// TIA Portal project "Est_clasificacion" (V17)

(* hardware
DEVICE "Estación S7-1500/ET200MP_1"  S7-1500 station
   slot 0: "Perfil soporte_0"  Rack  6ES7 590-1***0-0AA0
   slot 1: "PLC_1"  CPU 1516-3 PN/DP  6ES7 516-3AN02-0AB0  V2.9
      slot 3: "Display de la CPU_1"  6ES7591-1BA00-0AA0
      slot 32768: "Interfaz PROFINET_1"  X1
         slot 32769: "Puerto_1"  X1 P1
         slot 32770: "Puerto_2"  X1 P2
      slot 33024: "Interfaz PROFINET_2"  X2
         slot 33025: "Puerto_1"  X2 P1
      slot 33280: "Interfaz DP_1"  X3
      slot 34817: "Virtual CP interface port_1"  Virtual CP interface port  Virtual CP interface port
   slot 2: "DI 32x24VDC HF_1"  DI 32x24VDC HF  6ES7 521-1BL00-0AB0  V2.2
   slot 3: "DQ 32x24VDC/0.5A HF_1"  DQ 32x24VDC/0.5A HF  6ES7 522-1BL01-0AB0  V1.1
   slot 4: "AI 8xU/I/RTD/TC ST_1"  AI 8xU/I/RTD/TC ST  6ES7 531-7KF00-0AB0  V2.2
   slot 5: "AQ 4xU/I ST_1"  AQ 4xU/I ST  6ES7 532-5HD00-0AB0  V2.2
DEVICE "HMI_1"  KTP600 Basic color PN
   slot 0: "HMI_1"  KTP600 Basic color PN  6AV6 647-0AD11-3AX0  12.0.0.0
   slot 1: "HMI_RT_1"  KTP600 Basic color PN  6AV6 647-0AD11-3AX0  12.0.0.0
   slot 5: "HMI_1.IE_CP_1"  PROFINET Interface  12.0.0.0
      slot 1: "Interfaz PROFINET_1"  PROFINET Interface
         slot 1: "Port_1"  Port
*)

// ===== PLC "PLC_1"  CPU 1516-3 PN/DP =====

VAR_GLOBAL   // PLC tag table "Tabla de variables estándar"
   "Detector pieza inicio" AT %I0.0 : Bool;
   "Deflector 1" AT %I0.1 : Bool;
   "Detector de pieza" AT %I0.2 : Bool;
   "Deflector 2" AT %I0.3 : Bool;
   "Detector pieza color" AT %I0.4 : Bool;
   "Detector pieza negra" AT %I0.5 : Bool;
   "Detector pieza metalica" AT %I0.6 : Bool;
   "Start" AT %I1.0 : Bool;
   "Reset" AT %I1.3 : Bool;
   "Avanzar cinta" AT %Q0.0 : Bool;
   "Avanzar deflector 1" AT %Q0.1 : Bool;
   "Avanzar deflector 2" AT %Q0.2 : Bool;
   "Retraer tope" AT %Q0.3 : Bool;
   "Luz ON" AT %Q1.0 : Bool;
   "Luz RESET" AT %Q1.1 : Bool;
   "M0.0" AT %M0.0 : Bool;
   "M0.1" AT %M0.1 : Bool;
   "M0.2" AT %M0.2 : Bool;
   "C0.0" AT %M0.3 : Bool;
   "C0.1" AT %M0.4 : Bool;
   "C0.2" AT %M0.5 : Bool;
   "M1.0" AT %M1.0 : Bool;
   "M1.1" AT %M1.1 : Bool;
   "M1.2" AT %M1.2 : Bool;
   "M1.3" AT %M1.3 : Bool;
   "M1.4" AT %M1.4 : Bool;
   "M1.5" AT %M1.5 : Bool;
   "System_Byte" AT %MB7789 : Byte;
   "FirstScan" AT %M7789.0 : Bool;
   "DiagStatusUpdate" AT %M7789.1 : Bool;
   "AlwaysTRUE" AT %M7789.2 : Bool;
   "AlwaysFALSE" AT %M7789.3 : Bool;
END_VAR

// folder: System blocks/Program resources

DATA_BLOCK "IEC_Timer_0_DB"   // DB1
{ S7_Optimized_Access := 'TRUE' }
AUTHOR : Simatic
FAMILY : IEC
NAME : IEC_TMR
VERSION : 1.0
// stored: InstanceOfName IEC_TIMER
"IEC_TIMER"
BEGIN
END_DATA_BLOCK

DATA_BLOCK "IEC_Counter_0_DB"   // DB4
{ S7_Optimized_Access := 'TRUE' }
AUTHOR : Simatic
FAMILY : IEC
NAME : CNTR
VERSION : 1.0
// stored: InstanceOfName IEC_COUNTER
"IEC_COUNTER"
BEGIN
END_DATA_BLOCK

DATA_BLOCK "IEC_Counter_0_DB_1"   // DB5
{ S7_Optimized_Access := 'TRUE' }
AUTHOR : Simatic
FAMILY : IEC
NAME : CNTR
VERSION : 1.0
// stored: InstanceOfName IEC_COUNTER
"IEC_COUNTER"
BEGIN
END_DATA_BLOCK

DATA_BLOCK "IEC_Counter_0_DB_2"   // DB6
{ S7_Optimized_Access := 'TRUE' }
AUTHOR : Simatic
FAMILY : IEC
NAME : CNTR
VERSION : 1.0
// stored: InstanceOfName IEC_COUNTER
"IEC_COUNTER"
BEGIN
END_DATA_BLOCK

// folder: (top level)

ORGANIZATION_BLOCK "Main"   // OB1, LAD, ProgramCycle
TITLE = "Main Program Sweep (Cycle)"
{ S7_Optimized_Access := 'TRUE' }
VERSION : 0.1
   VAR_INPUT
      Initial_Call : Bool;   // Initial call of this OB
      Remanence : Bool;   // =True, if remanent data are available
   END_VAR
   VAR_TEMP   // added for the SCL form of the ladder/FBD networks
      _w1 : Bool;
      _w2 : Bool;
   END_VAR
BEGIN

REGION Network 1: Estados panel
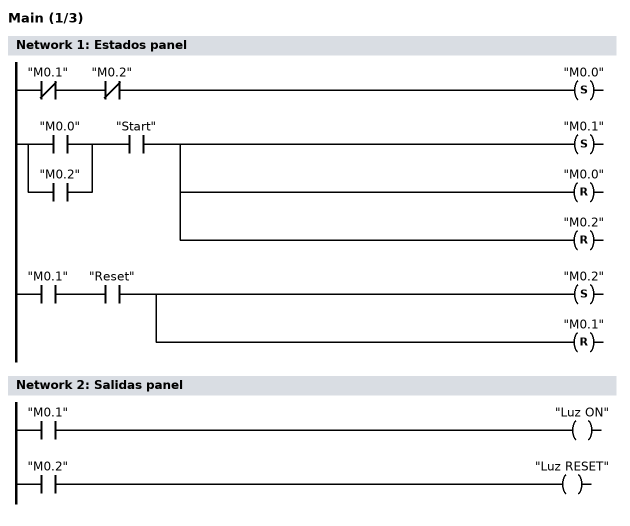
   RUNG wire#powerrail
      I_Contact( "M0.1" )
      I_Contact( "M0.2" )
      S_Coil( "M0.0" )
   END_RUNG
   RUNG wire#powerrail
      Contact( "M0.0" )
      wire#w1
      Contact( "Start" )
      wire#w2
      S_Coil( "M0.1" )
   END_RUNG
   RUNG wire#powerrail
      Contact( "M0.2" )
   END_RUNG wire#w1
   RUNG wire#w2
      R_Coil( "M0.0" )
   END_RUNG
   RUNG wire#w2
      R_Coil( "M0.2" )
   END_RUNG
   RUNG wire#powerrail
      Contact( "M0.1" )
      Contact( "Reset" )
      wire#w3
      S_Coil( "M0.2" )
   END_RUNG
   RUNG wire#w3
      R_Coil( "M0.1" )
   END_RUNG
   // the same network as SCL:
   IF NOT "M0.1" AND NOT "M0.2" THEN "M0.0" := TRUE; END_IF;
   IF ("M0.0" OR "M0.2") AND "Start" THEN "M0.1" := TRUE; END_IF;
   #_w1 := ("M0.0" OR "M0.2") AND "Start";
   IF #_w1 THEN
       "M0.0" := FALSE;
       "M0.2" := FALSE;
   END_IF;
   IF "M0.1" AND "Reset" THEN
       "M0.2" := TRUE;
       "M0.1" := FALSE;
   END_IF;
END_REGION

REGION Network 2: Salidas panel
   RUNG wire#powerrail
      Contact( "M0.1" )
      Coil( "Luz ON" )
   END_RUNG
   RUNG wire#powerrail
      Contact( "M0.2" )
      Coil( "Luz RESET" )
   END_RUNG
   // the same network as SCL:
   "Luz ON" := "M0.1";
   "Luz RESET" := "M0.2";
END_REGION

REGION Network 3: Estados principal
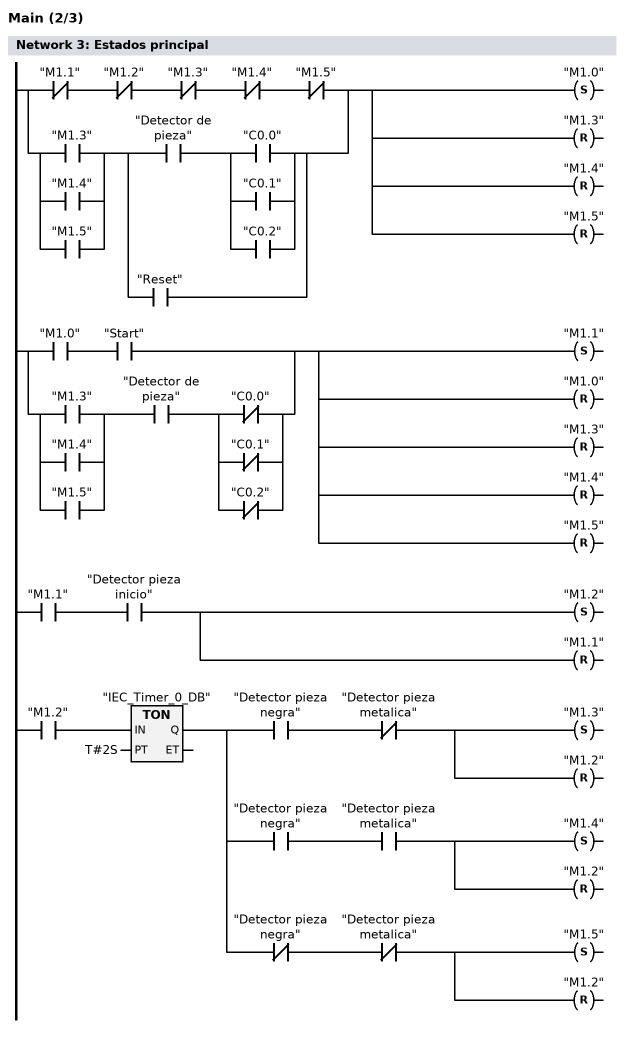
   IF (NOT "M1.1" AND NOT "M1.2" AND NOT "M1.3" AND NOT "M1.4" AND NOT "M1.5") OR (("M1.3" OR "M1.4" OR "M1.5") AND (("Detector de pieza" AND ("C0.0" OR "C0.1" OR "C0.2")) OR "Reset")) THEN
       "M1.0" := TRUE;
   END_IF;
   #_w1 := (NOT "M1.1" AND NOT "M1.2" AND NOT "M1.3" AND NOT "M1.4" AND NOT "M1.5") OR (("M1.3" OR "M1.4" OR "M1.5") AND (("Detector de pieza" AND ("C0.0" OR "C0.1" OR "C0.2")) OR "Reset"));
   IF #_w1 THEN
       "M1.3" := FALSE;
       "M1.4" := FALSE;
       "M1.5" := FALSE;
   END_IF;
   IF ("M1.0" AND "Start") OR (("M1.3" OR "M1.4" OR "M1.5") AND "Detector de pieza" AND (NOT "C0.0" OR NOT "C0.1" OR NOT "C0.2")) THEN
       "M1.1" := TRUE;
   END_IF;
   #_w2 := ("M1.0" AND "Start") OR (("M1.3" OR "M1.4" OR "M1.5") AND "Detector de pieza" AND (NOT "C0.0" OR NOT "C0.1" OR NOT "C0.2"));
   IF #_w2 THEN
       "M1.0" := FALSE;
       "M1.3" := FALSE;
       "M1.4" := FALSE;
       "M1.5" := FALSE;
   END_IF;
   IF "M1.1" AND "Detector pieza inicio" THEN
       "M1.2" := TRUE;
       "M1.1" := FALSE;
   END_IF;
   "IEC_Timer_0_DB".TON(IN := "M1.2", PT := T#2S);
   IF "IEC_Timer_0_DB".Q AND "Detector pieza negra" AND NOT "Detector pieza metalica" THEN
       "M1.3" := TRUE;
       "M1.2" := FALSE;
   END_IF;
   IF "IEC_Timer_0_DB".Q AND "Detector pieza negra" AND "Detector pieza metalica" THEN
       "M1.4" := TRUE;
       "M1.2" := FALSE;
   END_IF;
   IF "IEC_Timer_0_DB".Q AND NOT "Detector pieza negra" AND NOT "Detector pieza metalica" THEN
       "M1.5" := TRUE;
       "M1.2" := FALSE;
   END_IF;
END_REGION

REGION Network 4: Salidas principal
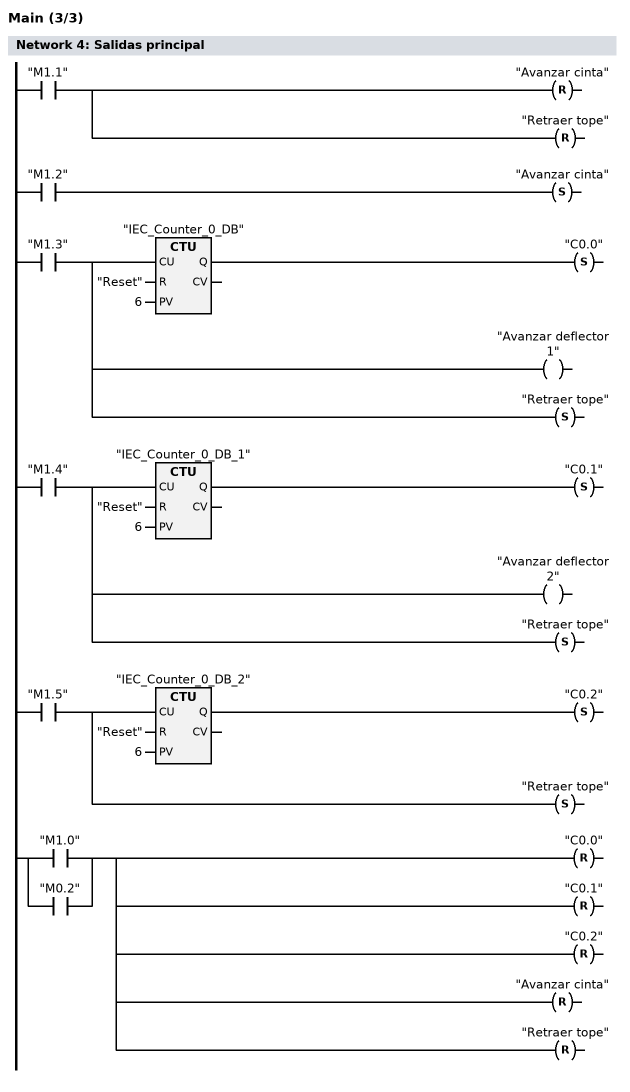
   IF "M1.1" THEN
       "Avanzar cinta" := FALSE;
       "Retraer tope" := FALSE;
   END_IF;
   IF "M1.2" THEN "Avanzar cinta" := TRUE; END_IF;
   "IEC_Counter_0_DB".CTU(CU := "M1.3", R := "Reset", PV := 6);
   IF "IEC_Counter_0_DB".Q THEN "C0.0" := TRUE; END_IF;
   "Avanzar deflector 1" := "M1.3";
   IF "M1.3" THEN "Retraer tope" := TRUE; END_IF;
   "IEC_Counter_0_DB_1".CTU(CU := "M1.4", R := "Reset", PV := 6);
   IF "IEC_Counter_0_DB_1".Q THEN "C0.1" := TRUE; END_IF;
   "Avanzar deflector 2" := "M1.4";
   IF "M1.4" THEN "Retraer tope" := TRUE; END_IF;
   "IEC_Counter_0_DB_2".CTU(CU := "M1.5", R := "Reset", PV := 6);
   IF "IEC_Counter_0_DB_2".Q THEN "C0.2" := TRUE; END_IF;
   IF "M1.5" THEN "Retraer tope" := TRUE; END_IF;
   IF "M1.0" OR "M0.2" THEN
       "C0.0" := FALSE;
       "C0.1" := FALSE;
       "C0.2" := FALSE;
       "Avanzar cinta" := FALSE;
       "Retraer tope" := FALSE;
   END_IF;
END_REGION
END_ORGANIZATION_BLOCK

ORGANIZATION_BLOCK "Startup"   // OB100, LAD, Startup
TITLE = "Complete Restart"
{ S7_Optimized_Access := 'TRUE' }
VERSION : 0.1
   VAR_INPUT
      LostRetentive : Bool;   // True if retentive data are lost
      LostRTC : Bool;   // True if date and time are lost
   END_VAR
BEGIN

REGION Network 1
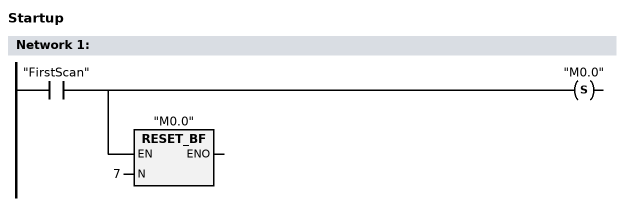
   // no SCL statement known for RBitfield: written as a call
   IF "FirstScan" THEN
       "M0.0" := TRUE;
       RESET_BF(operand := "M0.0", n := 7);
   END_IF;
END_REGION
END_ORGANIZATION_BLOCK

(* ===== HMI "HMI_RT_1" =====
system functions are stored by id; their names below are inferred from use
connection "HMI_Conexión_1": ETHERNET, SMART_S7_1500_OMS

HMI tags "Tabla de variables estándar"
   "Número_imagen_variable" : UInt, internal
   "Start" : Bool = PLC Start AT %I1.0, 1 s
   "Reset" : Bool = PLC Reset AT %I1.3, 1 s
   "C0.0" : Bool = PLC "C0.0" AT %M0.3, 1 s
   "IEC_Counter_0_DB_CV" : Int = PLC IEC_Counter_0_DB.CV, 1 s
   "IEC_Counter_0_DB_1_CV" : Int = PLC IEC_Counter_0_DB_1.CV, 1 s
   "IEC_Counter_0_DB_2_CV" : Int = PLC IEC_Counter_0_DB_2.CV, 1 s

text list "Nombre_imagen_lista_texto": 1 'Imagen raíz'; 2 'Control'; 3 'Imágenes de sistema'; 4 'Información de sistema'

Template "Plantilla_1" 320x240
   Button "Salir" at 266,202 size 52x37; TextOff 'Salir'; PictureOff "ExitRuntime_KTP600_Basic_color_PN"; PictureOn "ExitRuntime_KTP600_Basic_color_PN"
      on Release: StopRuntime(0)
   Button "Template_Button" at 213,202 size 52x37; TextOff 'Text'
   Button "Template_Button_1" at 160,202 size 52x37; TextOff 'Text'
   Button "Template_Button_2" at 107,202 size 52x37; TextOff 'Text'
   Button "Template_Button_3" at 54,202 size 52x37; TextOff 'Control'
      on Press: ActivateScreen("Control", 0)
   Button "Imagen inicial" at 1,202 size 52x37; TextOff 'Imagen inicial'; PictureOff "NavigateHome_KTP600_Basic_color_PN"; PictureOn "NavigateHome_KTP600_Basic_color_PN"
      on Release: ActivateScreen("Imagen raíz", 0)
   SymbolicIOField "Imagen_campo_ES_simbólico" at 59,7 size 259x24; TextOff '0'; TextOn '1'; TextList "Nombre_imagen_lista_texto"
      ProcessValue <- "Número_imagen_variable"
      on Change: ActivateScreenByNumber("Número_imagen_variable", 0)
   GraphicView "Logotipo" at 0,0 size 57x38; Picture "Logotipo de HMI_1"

screen "Imagen raíz" 320x240, template "Plantilla_1"
   on GenerateScreen: SetTag("Número_imagen_variable", 1)
   TextField "HmiScreenItemData" at 29,45 size 256x17; Text 'Bienvenido a la estacion de clasificacion!'
   GraphicView "Visor de gráficos_1" at 94,73 size 130x112; Picture "Gráfico_2"

screen "Control" 320x240, template "Plantilla_1"
   on GenerateScreen: SetTag("Número_imagen_variable", 2)
   Button "Botón_1" at 27,71 size 96x32; TextOff 'ON'
      on Press: SetBit("Start")
   Button "Botón_2" at 27,127 size 96x32; TextOff 'Reset'
      on Press: SetBit("Reset")
   TextField "Campo de texto_1" at 243,71 size 10x13; Text '0'
      Visibility <- "IEC_Counter_0_DB_CV"
   TextField "Campo de texto_2" at 202,69 size 35x15; Text 'ROJO:'
   TextField "Campo de texto_3" at 254,117 size 10x13; Text '0'
      Visibility <- "IEC_Counter_0_DB_1_CV"
   TextField "Campo de texto_4" at 202,114 size 42x16; Text 'PLATA'
   TextField "Campo de texto_5" at 253,155 size 10x13; Text '0'
      Visibility <- "IEC_Counter_0_DB_2_CV"
   TextField "Campo de texto_6" at 198,153 size 39x15; Text 'NEGRO'

screen "Imágenes de sistema" 320x240, template "Plantilla_1"
   on GenerateScreen: SetTag("Número_imagen_variable", 3)
   TextField "HmiScreenItemData" at 32,109 size 256x17; Text 'Imágenes de sistema'
   Button "Atrás" at 1,39 size 104x30; TextOff 'Atrás'
      on Release: ActivateScreen("Imagen raíz", 0)
   Button "Información de sistema" at 106,39 size 104x30; TextOff 'Información de ...'
      on Release: ActivateScreen("Información de sistema", 0)

screen "Información de sistema" 320x240, template "Plantilla_1"
   on GenerateScreen: SetTag("Número_imagen_variable", 4)
   TextField "HmiScreenItemData" at 4,71 size 120x20; Text 'Tipo de panel:'
   TextField "HmiScreenItemData_1" at 128,71 size 188x20; Text 'KTP600 Basic color PN 12.0'
   TextField "HmiScreenItemData_2" at 4,92 size 120x20; Text 'Conexión:'
   TextField "HmiScreenItemData_3" at 128,92 size 188x20; Text 'PROFINET (X1)'
   TextField "HmiScreenItemData_4" at 4,113 size 120x20; Text 'Controlador:'
   TextField "HmiScreenItemData_5" at 128,113 size 188x20; Text 'SIMATIC S7 1500'
   Button "Atrás" at 1,39 size 104x30; TextOff 'Atrás'
      on Release: ActivateScreen("Imágenes de sistema", 0)
*)